
   // BODY (data max. 232 Byte, Array 0..231 of Byte) 
   IF #RD_WR = TRUE THEN
       // IO-Link write data record requested, copy data from "RECORD_IOL_DATA"
       #write.header.IOL.Control := B#16#02; // CONTROL B#16#02 = write data record
       #wrrec.length := INT_TO_UINT(#LEN) + UINT#8;  // data length header + data = IO-Link write data record
       #typeofrequest := 2; // write data record
       // copy IOL_RECORD_DATA in working area
       #i := INT#0;    // initialize loop counter 
       FOR #i := 0 TO #LEN - 1 DO
           #write.data[#i] := #RECORD_IOL_DATA[#i];
       END_FOR;
   ELSE
       // IO-Link read data record requested
       #write.header.IOL.Control := 16#03;  // CONTROL 16#03 = read data record
       #wrrec.length := UINT#8; // data length only header = IO-Link read data record
       #typeofrequest := 1; // read data record        
   END_IF;
   #sequencecontrol := 1;  // Start sequence
   ELSE
       ;
   END_IF;

   (*---------------------------------------------------------------------------------------------------------------------
               SEQUENCE CONTROL
   ---------------------------------------------------------------------------------------------------------------------*)
   CASE #sequencecontrol OF
       1:  // Check input parameter        
           IF #PORT < INT#0 OR #PORT > INT#63 THEN // PORT (Wrong port address = 0x8001)
               #ERROR := TRUE;
               #IOL_STATUS := DW#16#80010000;
               #sequencecontrol := 99; // aborting function with error
           ELSIF #IOL_INDEX < INT#0 OR #IOL_INDEX > INT#32767 THEN    // INDEX (Wrong index = 0x8002)
               #ERROR := TRUE;
               #IOL_STATUS := DW#16#80020000;
               #sequencecontrol := 99; // aborting function with error
           ELSIF #IOL_SUBINDEX < INT#0 OR #IOL_SUBINDEX > INT#255 THEN    // SUBINDEX (Wrong subindex = 0x8003)
               #ERROR := TRUE;
               #IOL_STATUS := DW#16#80030000;
               #sequencecontrol := 99; // aborting function with error
           ELSIF #typeofrequest = 2 AND (#LEN < 1 OR #LEN > 232) THEN  // LEN (wrong length for write data record = 0x8004)
               #ERROR := TRUE;
               #IOL_STATUS := DW#16#80050000;
               #sequencecontrol := 99; // aborting function with error
           ELSIF #typeofrequest = 1 AND (#LEN < 0 OR #LEN > 232) THEN  // LEN (wrong length for read data record = 0x8005)
               #ERROR := TRUE;
               #IOL_STATUS := DW#16#80060000;
               #sequencecontrol := 99; // aborting function with error
           ELSE    // all input parameter are right
               #sequencecontrol := 2;
           END_IF;

       2:  (*-------------------------------------------------------------------------------------------------------------
           WRREC = Write Data Record
           Note:
           To read data records, the IO-Link master modules needs to know which PORT is required. Therefore it is necessary
           to send at first a request via write data record (header, 8 byte). As response the IO-Link master module will 
           send the required data record.
           -------------------------------------------------------------------------------------------------------------*)
           #WRREC_Function(REQ := TRUE,
                           LEN := #wrrec.length,
                           DONE => #wrrec.done,
                           BUSY => #wrrec.busy,
                           ERROR => #wrrec.error,
                           STATUS => #wrrec.status,
                           RECORD := #write);
           // output status during write data record
           IF #wrrec.busy THEN
               #STATUS := #wrrec.status;
               #IOL_STATUS := DW#16#00020000;  // 0002 = writing in progress 
           ELSIF #wrrec.error THEN
               #tmpDWORD := #wrrec.status AND DW#16#00FFFF00;  // filter status
               IF #tmpDWORD = DW#16#0080C200 THEN    // if resource #BUSY (#STATUS=80C2), then ... 
                   #sequencecontrol := 3;  // ... repeat write data record
               ELSE
                   #ERROR := TRUE;
                   #STATUS := #wrrec.status;   // ... otherwise output error status of "WRREC"
                   #IOL_STATUS := DW#16#80530000;  // ... with note '8053' = error status of "WRREC"
                   #sequencecontrol := 99; // aborting function with error
               END_IF;
           ELSIF #wrrec.done = TRUE THEN   // wait for write data record finish without error
               #TP_poll(IN := TRUE,
                        PT := T#100ms);    // poll for response
               #sequencecontrol := 4;
           ELSE
               ;
           END_IF;

       3:  // repeat write data record because resource was busy
           #WRREC_Function(REQ := FALSE);
           #sequencecontrol := 2;

       4:  // wait and poll for response = Read Data Record (RDREC)
           #WRREC_Function(REQ := FALSE);
           #TP_poll(IN := TRUE,
                    PT := T#100ms);

           // if poll rate executed then start read data record (on falling edge)
           #F_TRIG_poll := #TP_poll.Q = FALSE AND #F_TRIG_poll_old = TRUE;
           #F_TRIG_poll_old := #TP_poll.Q = TRUE;

           // RDREC = Read Data Record
           #RDREC_Function(REQ := #F_TRIG_poll,
                           MLEN := UINT#0, // length = 0 = read all data which are available
                           VALID => #rdrec.valid,
                           BUSY => #rdrec.busy,
                           ERROR => #rdrec.error,
                           STATUS => #rdrec.status,
                           LEN => #rdrec.length,
                           RECORD := #read);
           // output status during read data record
           IF #rdrec.busy THEN
               #STATUS := #rdrec.status;
               #IOL_STATUS := DW#16#00030000; // 16#0003 = reading in progress
           ELSIF #rdrec.error = TRUE THEN
               #tmpDWORD := #rdrec.status AND DW#16#00FFFF00;  // filter status
               IF #tmpDWORD = DW#16#0080C200 THEN  // if resource busy (status=80C2), then ... 
                   #sequencecontrol := 5;  // ... repeat read data record / continue polling
               ELSE
                   #ERROR := TRUE;
                   #STATUS := #rdrec.status;   // ... otherwise output error code of "RDREC"
                   #IOL_STATUS := DW#16#80520000;  // ... with note '8052' = error status of "RDREC"
                   #sequencecontrol := 99; // aborting function with error
               END_IF;
           ELSIF #rdrec.valid THEN
               IF  // check the response wether it matches the request (compare PORT, INDEX and SUBINDEX)
                   (#write.header.CALL.Port <> #read.header.CALL.Port) OR
                   (#write.header.IOL.Index_HighByte <> #read.header.IOL.Index_HighByte) OR
                   (#write.header.IOL.Index_LowByte <> #read.header.IOL.Index_LowByte) OR
                   (#write.header.IOL.Subindex <> #read.header.IOL.Subindex)
               THEN    // read data record don't match the request
                   #ERROR := TRUE;
                   #STATUS := #rdrec.status;
                   #IOL_STATUS := DW#16#70000000;  // output status '7000', no consistent data
                   #sequencecontrol := 99; // aborting function with error
               ELSIF #read.header.IOL.Control = B#16#80 THEN   // check the response for IO-Link errors
                   // State 0x80 = IOL_CALL_RES PDU shows IO-Link error detect
                   #ERROR := TRUE;
                   #STATUS := DW#16#00000000;
                   #IOL_STATUS.%B3 := #read.data[0];   // IO-Link master error code
                   #IOL_STATUS.%B2 := #read.data[1];   // IO-Link master error code
                   #IOL_STATUS.%B1 := #read.data[2];  // IO-Link device error code
                   #IOL_STATUS.%B0 := #read.data[3];  // IO-Link device additional error code

                   #sequencecontrol := 99; // aborting function with error
               ELSE    // read data are valid = output
                   #DONE_VALID := TRUE;
                   #BUSY := FALSE;
                   #ERROR := FALSE;
                   #STATUS := DW#16#00000000;
                   #IOL_STATUS := DW#16#00000000;  // request finished

                   IF #typeofrequest = 1 THEN
                       #RD_LEN := UINT_TO_INT(#rdrec.length - UINT#8);  // device parameter cover header and data,
                       // only data will be output
                       #i := INT#0; // initialize loop counter
                       FOR #i := 0 TO UINT_TO_INT(#rdrec.length - UINT#8 - UINT#1) DO
                           #RECORD_IOL_DATA[#i] := #read.data[#i];
                       END_FOR;
                   ELSE
                       ;
                   END_IF;
                   #sequencecontrol := 98;
               END_IF;
           ELSE
               ;
           END_IF;

       5:  // poll again for response because resource was busy
           #TP_poll(IN := FALSE,
                    PT := T#100ms);
           #RDREC_Function(REQ := FALSE,
                           RECORD := #read);
           #sequencecontrol := 4;  // ... repeat read data record / continue polling   

       98: // request done successfully
           #TP_poll(IN := FALSE,
                    PT := T#100ms);
           #RDREC_Function(REQ := FALSE,
                           RECORD := #read);
           IF #REQ = FALSE THEN
               #DONE_VALID := FALSE;
               #BUSY := FALSE;
               #ERROR := FALSE;
               #RD_LEN := INT#0;
               #STATUS := DW#16#00000000;
               #IOL_STATUS := DW#16#00010000; // ready for new request
               #sequencecontrol := 0;
               #typeofrequest := 0;
           ELSE
               ;
           END_IF;

       99: // Function aborted with error
           #TP_poll(IN := FALSE,
                    PT := T#100ms);
           #WRREC_Function(REQ := FALSE);
           #RDREC_Function(REQ := FALSE,
                           RECORD := #read);
           #DONE_VALID := FALSE;
           #BUSY := FALSE;
           #RD_LEN := INT#0;
           #sequencecontrol := 0;
           #typeofrequest := 0;

       ELSE  // no relevant case, ready for new request
           #WRREC_Function(REQ := FALSE);
           #RDREC_Function(REQ := FALSE,
                           RECORD := #read);
           #TP_poll(IN := FALSE,
                    PT := T#100ms);
           #TON_monitoring(IN := FALSE,
                           PT := T#20s);
           #sequencecontrol := 0;
           #typeofrequest := 0;
   END_CASE;

   (*---------------------------------------------------------------------------------------------------------------------
               MONITORING
   ---------------------------------------------------------------------------------------------------------------------*)
   #TON_monitoring(IN := #sequencecontrol > 0 AND #sequencecontrol < 98,
                   PT := T#20s);
   IF #TON_monitoring.Q THEN
       #ERROR := TRUE;
       #IOL_STATUS := DW#16#80000000; // request time out       
       #sequencecontrol := 99; // aborting function with error
   END_IF;
END_FUNCTION_BLOCK

(* ===== HMI "HMI_RT_1" =====
system functions are stored by id; their names below are inferred from use
connection "HMI_Connection_1": ETHERNET, SMART_S7_1200_OMS

HMI tags "Default tag table"
   "Emergency Stop Stacker" : Bool = PLC 113S1 AT %I1.0, 1 s
   "Avarie Conveior 4 stacker" : Bool = PLC 128U1_Fault AT %I5.1, 1 s
   "Prezenta aer" : Bool = PLC 151S1 AT %I2.0, 1 s
   "Protectie cuplata Conveior 1 alimentare destacker" : Bool = PLC 120Q1 AT %I2.2, 1 s
   "Protectie cuplata Conveior 2 iesire destacker" : Bool = PLC 122Q1 AT %I2.7, 1 s
   "Avarie Conveior 1 alimentare destacker" : Bool = PLC 120U1_Fault AT %I2.6, 1 s
   "Avarie Conveior 2 iesire destacker" : Bool = PLC 122U1_Fault AT %I3.3, 1 s
   "Contactor cuplat Conveior 1 alimentare destacker" : Bool = PLC 121K1 AT %I2.3, 1 s
   "Contactor cuplat Conveior 2 iesire destacker" : Bool = PLC 123K1 AT %I3.0, 1 s
   "Frana decuplata Conveior 1 alimentare destacker" : Bool = PLC 120K1 AT %I2.4, 1 s
   "Frana decuplata Conveior 2 iesire destacker" : Bool = PLC 122K1 AT %I3.1, 1 s
   "Functionare Conveior 1 alimentare destacker" : Bool = PLC 120U1_PowerOK AT %I2.5, 1 s
   "Functionare Conveior 2 iesire destacker" : Bool = PLC 122U1_PowerOK AT %I3.2, 1 s
   "Senzor 1 proximitate softstarter aer destacker" : Bool = PLC 142VFA1_SQ1 AT %I6.4, 1 s
   "Senzor 2 proximitate softstarter aer destacker" : Bool = PLC 142VFA1_SQ2 AT %I6.5, 1 s
   "Reset safety Destacker" : Bool = PLC 1XXS2 AT %I68.6, 1 s
   "Comanda 1 softstarter aer destacker" : Bool = PLC "Comanda 1 softstarter aer stacker_new" AT %Q64.1, 1 s
   "Cuplare contactor VFD Conveior 1 alimentare destacker" : Bool = PLC CSN3_PowerOK AT %Q7.3, 1 s
   "Fault Aknowledge VFD Conveior 1 alimentare destacker" : Bool = PLC CSN3_FaultAck AT %Q10.0, 1 s
   "ON/OFF1 VFD Conveior 1 alimentare destacker" : Bool = PLC CSN3_Start AT %Q7.4, 1 s
   "Cuplare contactor VFD Conveior 2 iesire destacker" : Bool = PLC CSN4_PowerOK AT %Q7.5, 1 s
   "Fault Aknowledge VFD Conveior 2 iesire destacker" : Bool = PLC CSN4_FaultAck AT %Q10.1, 1 s
   "ON/OFF1 VFD Conveior 2 iesire destacker" : Bool = PLC CSN4_Start AT %Q7.6, 1 s
   "Contactor cuplat Conveior 4 descarcare stacker" : Bool = PLC 129K1 AT %I4.6, 1 s
   "Frana decuplata Conveior 4 descarcare stacker" : Bool = PLC 128K1 AT %I4.7, 1 s
   "Functionare Conveior 4 stacker" : Bool = PLC 128U1_PowerOK AT %I5.0, 1 s
   "Protectie cuplata Conveior 4 descarcare stacker" : Bool = PLC 128Q1 AT %I4.5, 1 s
   "Cuplare contactor VFD Conveior 4 descarcare stacker" : Bool = PLC CS4_PowerOK AT %Q8.5, 1 s
   "Fault Aknowledge VFD Conveior 4 descarcare stacker" : Bool = PLC CS4_FaultAck AT %Q10.3, 1 s
   "ON/OFF1 VFD Conveior 4 descarcare stacker" : Bool = PLC CS4_Start AT %Q8.6, 1 s
   "Avarie Conveior 3 transfer palet 2" : Bool = PLC 126U1_Fault AT %I4.4, 1 s
   "Contactor cuplat Conveior 3 transfer palet 2" : Bool = PLC 127K1 AT %I4.1, 1 s
   "Frana decuplata Conveior 3 transfer palet 2" : Bool = PLC 126K1 AT %I4.2, 1 s
   "Functionare Conveior 1 preluare paleti OK" : Bool = PLC 124K1 AT %I3.5, 1 s
   "Functionare Conveior 2 transfer palet 1" : Bool = PLC 125K1 AT %I3.7, 1 s
   "Functionare Conveior 3 transfer palet 2" : Bool = PLC 126U1_PowerOK AT %I4.3, 1 s
   "Protectie cuplata Conveior 1 preluare paleti OK" : Bool = PLC 124Q1 AT %I3.4, 1 s
   "Protectie cuplata Conveior 2 transfer palet 1" : Bool = PLC 125Q1 AT %I3.6, 1 s
   "Protectie cuplata Conveior 3 transfer palet 2" : Bool = PLC 126Q1 AT %I4.0, 1 s
   "Cuplare contactor VFD Conveior 3 transfer palet 2" : Bool = PLC CS3_PowerOK AT %Q8.3, 1 s
   "Fault Aknowledge VFD Conveior 3 transfer palet 2" : Bool = PLC CS3_FaultAck AT %Q10.2, 1 s
   "ON/OFF1 VFD Conveior 3 transfer palet 2" : Bool = PLC CS3_Start AT %Q8.4, 1 s
   "Softstarter aer 1.1 Conveior 1 preluare paleti OK" : Bool = PLC "Softstarter aer 1.1 Conveior 1 preluare paleti OK" AT %Q8.1, 1 s
   "Softstarter aer 1.2 Conveior 1 preluare paleti OK" : Bool = PLC "Softstarter aer 1.2 Conveior 1 preluare paleti OK" AT %Q8.2, 1 s
   "Start Conveior 1 preluare paleti OK" : Bool = PLC CS1_Start AT %Q8.0, 1 s
   "Start Conveior 2 transfer palet 1" : Bool = PLC CS2_Start AT %Q7.0, 1 s
   "Comanda 2 softstarter aer destacker" : Bool = PLC "Comanda 2 softstarter aer stacker_new" AT %Q66.1, 1 s
   "Comanda 1 softstarter aer stacker" : Bool = PLC "Comanda 1 softstarter aer stacker" AT %Q72.1, 1 s
   "Comanda 2 softstarter aer stacker" : Bool = PLC "Comanda 2 softstarter aer stacker" AT %Q74.1, 1 s
   "MD_IS1_SC_X1.0" : Bool = PLC "MD_IS1_SC_X1.0" AT %I70.0, 1 s
   "MD_IS1_SC_X1.1" : Bool = PLC "MD_IS1_SC_X1.1" AT %I70.1, 1 s
   "MD_IS1_SC_X1.2" : Bool = PLC "MD_IS1_SC_X1.2" AT %I70.2, 1 s
   "MD_IS1_SC_X1.3" : Bool = PLC "MD_IS1_SC_X1.3" AT %I70.3, 1 s
   "MD_IS1_SC_X1.4" : Bool = PLC "MD_IS1_SC_X1.4" AT %I70.4, 1 s
   "MD_IS1_SC_X1.5" : Bool = PLC "MD_IS1_SC_X1.5" AT %I70.5, 1 s
   "MD_IS1_SC_X1.6" : Bool = PLC "MD_IS1_SC_X1.6" AT %I70.6, 1 s
   "MD_IS1_SC_X1.7" : Bool = PLC "MD_IS1_SC_X1.7" AT %I70.7, 1 s
   "MD_IS2_SC_X1.0" : Bool = PLC "MD_IS2_SC_X1.0" AT %I75.0, 1 s
   "MD_IS2_SC_X1.1" : Bool = PLC "MD_IS2_SC_X1.1" AT %I75.1, 1 s
   "MD_IS2_SC_X1.2" : Bool = PLC "MD_IS2_SC_X1.2" AT %I75.2, 1 s
   "MD_IS2_SC_X1.3" : Bool = PLC "MD_IS2_SC_X1.3" AT %I75.3, 1 s
   "MD_IS2_SC_X1.4" : Bool = PLC "MD_IS2_SC_X1.4" AT %I75.4, 1 s
   "MD_IS2_SC_X1.5" : Bool = PLC "MD_IS2_SC_X1.5" AT %I75.5, 1 s
   "MD_IS2_SC_X1.6" : Bool = PLC "MD_IS2_SC_X1.6" AT %I75.6, 1 s
   "MD_IS2_SC_X1.7" : Bool = PLC "MD_IS2_SC_X1.7" AT %I75.7, 1 s
   "MD_OS_SC_X1.0" : Bool = PLC "MD_OS_SC_X1.0" AT %I92.0, 1 s
   "MD_OS_SC_X1.1" : Bool = PLC "MD_OS_SC_X1.1" AT %I93.0, 1 s
   "MD_OS_SC_X1.2" : Bool = PLC "MD_OS_SC_X1.2" AT %I92.1, 1 s
   "MD_OS_SC_X1.3" : Bool = PLC "MD_OS_SC_X1.3" AT %I93.1, 1 s
   "MD_OS_SC_X1.4" : Bool = PLC "MD_OS_SC_X1.4" AT %I92.2, 1 s
   "MD_OS_SC_X1.5" : Bool = PLC "MD_OS_SC_X1.5" AT %I93.2, 1 s
   "MS_IS1_SC_X1.0" : Bool = PLC "MS_IS1_SC_X1.0" AT %I80.0, 1 s
   "MS_IS1_SC_X1.1" : Bool = PLC "MS_IS1_SC_X1.1" AT %I80.1, 1 s
   "MS_IS1_SC_X1.2" : Bool = PLC "MS_IS1_SC_X1.2" AT %I80.2, 1 s
   "MS_IS1_SC_X1.3" : Bool = PLC "MS_IS1_SC_X1.3" AT %I80.3, 1 s
   "MS_IS1_SC_X1.4" : Bool = PLC "MS_IS1_SC_X1.4" AT %I80.4, 1 s
   "MS_IS1_SC_X1.5" : Bool = PLC "MS_IS1_SC_X1.5" AT %I80.5, 1 s
   "MS_IS1_SC_X1.6" : Bool = PLC "MS_IS1_SC_X1.6" AT %I80.6, 1 s
   "MS_IS1_SC_X1.7" : Bool = PLC "MS_IS1_SC_X1.7" AT %I80.7, 1 s
   "MS_IS2_SC_X1.0" : Bool = PLC "MS_IS2_SC_X1.0" AT %I85.0, 1 s
   "MS_IS2_SC_X1.1" : Bool = PLC "MS_IS2_SC_X1.1" AT %I85.1, 1 s
   "MS_IS2_SC_X1.2" : Bool = PLC "MS_IS2_SC_X1.2" AT %I85.2, 1 s
   "MS_IS2_SC_X1.3" : Bool = PLC "MS_IS2_SC_X1.3" AT %I85.3, 1 s
   "MS_IS2_SC_X1.4" : Bool = PLC "MS_IS2_SC_X1.4" AT %I85.4, 1 s
   "MS_IS2_SC_X1.5" : Bool = PLC "MS_IS2_SC_X1.5" AT %I85.5, 1 s
   "MS_IS2_SC_X1.6" : Bool = PLC "MS_IS2_SC_X1.6" AT %I85.6, 1 s
   "MS_IS2_SC_X1.7" : Bool = PLC "MS_IS2_SC_X1.7" AT %I85.7, 1 s
   "MS_OS_SC_X1.0" : Bool = PLC "MS_OS_SC_X1.0" AT %I101.0, 1 s
   "MS_OS_SC_X1.1" : Bool = PLC "MS_OS_SC_X1.1" AT %I102.0, 1 s
   "MS_OS_SC_X1.2" : Bool = PLC "MS_OS_SC_X1.2" AT %I101.1, 1 s
   "MS_OS_SC_X1.3" : Bool = PLC "MS_OS_SC_X1.3" AT %I102.1, 1 s
   "MS_OS_SC_X1.4" : Bool = PLC "MS_OS_SC_X1.4" AT %I101.2, 1 s
   "MS_OS_SC_X1.5" : Bool = PLC "MS_OS_SC_X1.5" AT %I102.2, 1 s
   "DS_Comanda cilindru vertical jos" : Bool = PLC "SN_Comanda cilindru vertical jos" AT %Q66.0, 1 s
   "DS_Comanda cilindru vertical sus" : Bool = PLC "SN_Comanda cilindru vertical sus" AT %Q64.0, 1 s
   "DS_Comanda furca retrasa" : Bool = PLC "SN_Comanda furca retrasa" AT %Q65.0, 1 s
   "DB_PalletDispenser_PD2_De_Stacking_DB_PD1_MiddlePosition" : Bool = PLC DB_PalletDispenser_PD2_Stacking_New_DB.PD1.MiddlePosition, 1 s
   "DB_PalletDispenser_PD2_De_Stacking_DB_PD1_Up" : Bool = PLC DB_PalletDispenser_PD2_Stacking_New_DB.PD1.Up, 1 s
   "DB_PalletDispenser_PD2_De_Stacking_DB_PD1_Down" : Bool = PLC DB3_FAULTS.Alarm_Safety_S, 1 s
   "DB_PalletDispenser_PD2_De_Stacking_DB_PD1_Forks_In" : Bool = PLC DB3_FAULTS.Alarm_Safety_Z2, 1 s
   "DB_PalletDispenser_PD2_De_Stacking_DB_PD1_Forks_Out" : Bool = PLC DB_PalletDispenser_PD2_Stacking_New_DB.PD1.Forks_Out, 1 s
   "DB_PalletDispenser_PD2_De_Stacking_DB_Alarm_Active" : Bool = PLC DB3_FAULTS.Alarm_CD1, 1 s
   "DB_PalletDispenser_PD2_Stacking_DB_PD1_MiddlePosition" : Bool = PLC DB_PalletDispenser_PD2_Stacking_DB.PD1.MiddlePosition, 1 s
   "DB_PalletDispenser_PD2_Stacking_DB_PD1_Up" : Bool = PLC DB_PalletDispenser_PD2_Stacking_DB.PD1.Up, 1 s
   "DB_PalletDispenser_PD2_Stacking_DB_PD1_Down" : Bool = PLC DB_PalletDispenser_PD2_Stacking_DB.PD1.Down, 1 s
   "DB_PalletDispenser_PD2_Stacking_DB_PD1_Forks_In" : Bool = PLC DB_PalletDispenser_PD2_Stacking_DB.PD1.Forks_In, 1 s
   "DB_PalletDispenser_PD2_Stacking_DB_PD1_Forks_Out" : Bool = PLC DB_PalletDispenser_PD2_Stacking_DB.PD1.Forks_Out, 1 s
   "DB_PalletDispenser_PD2_Stacking_DB_Alarm_Active" : Bool = PLC DB_PalletDispenser_PD2_Stacking_DB.Alarm.Active, 1 s
   "S_Comanda cilindru vertical jos" : Bool = PLC "S_Comanda cilindru vertical jos" AT %Q74.0, 1 s
   "S_Comanda cilindru vertical sus" : Bool = PLC "S_Comanda cilindru vertical sus" AT %Q72.0, 1 s
   "S_Comanda furca retrasa" : Bool = PLC "S_Comanda furca retrasa" AT %Q73.0, 1 s
   "S_Comanda furca extinsa" : Bool = PLC "S_Comanda furca extinsa" AT %Q75.0, 1 s
   "Destacker 110KF1 Safety Relay" : Bool = PLC 110KF1 AT %I0.0, 1 s
   "Destacker 111KF1 Safety Barrier Relay" : Bool = PLC 111KF1 AT %I0.1, 1 s
   "Emergency Stop Destacker" : Bool = PLC 110S1 AT %I0.6, 1 s
   "Emergency Stop Zone 2" : Bool = PLC 112S1 AT %I0.7, 1 s
   "Stacker 113KF1 Safety Relay" : Bool = PLC 113KF1 AT %I0.3, 1 s
   "Stacker 114KF1 Safety Barrier Relay 1" : Bool = PLC 114KF1 AT %I0.4, 1 s
   "Stacker 115KF1 Safety Barrier Relay 2" : Bool = PLC 115KF1 AT %I0.5, 1 s
   "Zone 2 112KF1 Safety Relay" : Bool = PLC 112KF1 AT %I0.2, 1 s
   "Reset Destacker 110KF1 Safety Relay" : Bool = PLC 153K1 AT %Q0.0, 1 s
   "Reset Destacker 111KF1 Safety Barrier Relay" : Bool = PLC 153K2 AT %Q0.1, 1 s
   "Reset safety Zone 2" : Bool = PLC 155S1 AT %I1.1, 1 s
   "Reset Stacker 113KF1 Safety Relay" : Bool = PLC 153K4 AT %Q0.3, 1 s
   "Reset Stacker 114KF1 Safety Barrier Relay 1" : Bool = PLC 153K5 AT %Q0.4, 1 s
   "Reset Stacker 115KF1 Safety Barrier Relay 2" : Bool = PLC 153K6 AT %Q0.5, 1 s
   "Reset Zone 2 112KF1 Safety Relay" : Bool = PLC 153K3 AT %Q0.2, 1 s
   "FB_AlarmCounter_DB_Counters_Destacker 110KF1 Safety Relay_CV" : Int = PLC FB_AlarmCounter_DB.Counters."Destacker 110KF1 Safety Relay".CV, 1 s
   "FB_AlarmCounter_DB_Counters_Destacker 111KF1 Safety Barrier Relay_CV" : Int = PLC FB_AlarmCounter_DB.Counters."Destacker 111KF1 Safety Barrier Relay".CV, 1 s
   "FB_AlarmCounter_DB_Counters_Zone 2 112KF1 Safety Relay_CV" : Int = PLC FB_AlarmCounter_DB.Counters."Zone 2 112KF1 Safety Relay".CV, 1 s
   "FB_AlarmCounter_DB_Counters_Stacker 113KF1 Safety Relay_CV" : Int = PLC FB_AlarmCounter_DB.Counters."Stacker 113KF1 Safety Relay".CV, 1 s
   "FB_AlarmCounter_DB_Counters_Stacker 114KF1 Safety Barrier Relay 1_CV" : Int = PLC FB_AlarmCounter_DB.Counters."Stacker 114KF1 Safety Barrier Relay 1".CV, 1 s
   "FB_AlarmCounter_DB_Counters_Stacker 115KF1 Safety Barrier Relay 2_CV" : Int = PLC FB_AlarmCounter_DB.Counters."Stacker 115KF1 Safety Barrier Relay 2".CV, 1 s
   "FB_AlarmCounter_DB_Counters_Emergency Stop Destacker_CV" : Int = PLC FB_AlarmCounter_DB.Counters."Emergency Stop Destacker".CV, 1 s
   "FB_AlarmCounter_DB_Counters_Emergency Stop Zone 2_CV" : Int = PLC FB_AlarmCounter_DB.Counters."Emergency Stop Zone 2".CV, 1 s
   "FB_AlarmCounter_DB_Counters_Emergency Stop Stacker_CV" : Int = PLC FB_AlarmCounter_DB.Counters."Emergency Stop Stacker".CV, 1 s
   "FB_EnergyCounter_DB_Counters_LastHour_CV" : UInt = PLC FB_EnergyCounter_DB.Counters.LastHour.CV, 1 s
   "FB_EnergyCounter_DB_Counters_LastDay_CV" : UDInt = PLC FB_EnergyCounter_DB.Counters.LastDay.CV, 1 s
   "FB_EnergyCounter_DB_Counters_LastMonth_CV" : UDInt = PLC FB_EnergyCounter_DB.Counters.LastMonth.CV, 1 s
   "Aliniere palet" : Bool = PLC CSN1_SQ3 AT %I68.1, 1 s
   "Centror extins" : Bool = PLC CP2_SQ3 AT %I79.5, 1 s
   "Centror retras" : Bool = PLC CP2_SQ2 AT %I78.5, 1 s
   "Detectie 1 aliniament palet" : Bool = PLC "Detectie 1 aliniament palet" AT %I69.1, 1 s
   "Detectie 2 aliniament palet" : Bool = PLC "Detectie 2 aliniament palet" AT %I68.2, 1 s
   "Detectie palet" : Bool = PLC "SN_Detectie palet" AT %I73.4, 1 s
   "DS_Cilindru extins" : Bool = PLC "SN_Cilindru extins" AT %I74.6, 1 s
   "DS_Cilindru retras" : Bool = PLC "SN_Cilindru retras" AT %I74.1, 1 s
   "DS_Cilindru vertical jos" : Bool = PLC "SN_Cilindru vertical jos" AT %I73.5, 1 s
   "DS_Cilindru vertical mijloc" : Bool = PLC "SN_Cilindru vertical mijloc" AT %I73.3, 1 s
   "DS_Cilindru vertical sus" : Bool = PLC "SN_Cilindru vertical sus" AT %I73.2, 1 s
   "DS_Lungime 1" : Bool = PLC CSN3_SQ2 AT %I68.3, 1 s
   "DS_Lungime 2" : Bool = PLC CSN3_SQ3 AT %I69.3, 1 s
   "DS_Lungime 3" : Bool = PLC CSN4_SQ1 AT %I68.4, 1 s
   "Feed palet" : Bool = PLC SN_Prez_conveyor_volum AT %I69.6, 1 s
   "Inaltime maxima" : Bool = PLC "Inaltime maxima" AT %I69.0, 1 s
   "Masurare lungime" : Bool = PLC CS2_SQ1 AT %I78.2, 1 s
   "Prezenta palet iesire" : Bool = PLC SN_Switch_Iesire AT %I69.4, 1 s
   "Prezenta palet_capat_conveyor" : Bool = PLC CS1_SQ3 AT %I78.1, 1 s
   "Prezenta palet_centror" : Bool = PLC "S_Prezenta palet_centror" AT %I79.1, 1 s
   "Prezenta palet_dreapta" : Bool = PLC "Prezenta palet_dreapta" AT %I79.0, 1 s
   "Prezenta palet_stanga" : Bool = PLC CS1_SQ1 AT %I78.0, 1 s
   "Prezenta_stiva" : Bool = PLC CS4_SQ1 AT %I78.4, 1 s
   "Prezenta stiva" : Bool = PLC CSN1_SQ1 AT %I68.0, 1 s
   "Protectie cuplata Circular masa fixa" : Bool = PLC 104F1 AT %I5.4, 1 s
   "Protectie cuplata HMI" : Bool = PLC 149F1 AT %I7.0, 1 s
   "Protectie cuplata Iluminat" : Bool = PLC 105F2 AT %I2.1, 1 s
   "Protectie cuplata Masina demontare paleti dreapta" : Bool = PLC 103F1 AT %I5.3, 1 s
   "Protectie cuplata Masina demontare paleti stanga" : Bool = PLC 102F1 AT %I5.2, 1 s
   "Protectie cuplata Post reparatie stanga+dreapta" : Bool = PLC 105F1 AT %I5.5, 1 s
   "Protectie cuplata Post reparatii minore" : Bool = PLC 106F1 AT %I5.6, 1 s
   "Protectie cuplata TELE" : Bool = PLC 107F1 AT %I5.7, 1 s
   "S_Cilindru extins" : Bool = PLC "S_Cilindru extins" AT %I84.6, 1 s
   "S_Cilindru retras" : Bool = PLC "S_Cilindru retras" AT %I84.1, 1 s
   "S_Cilindru vertical jos" : Bool = PLC "S_Cilindru vertical jos" AT %I83.5, 1 s
   "S_Cilindru vertical mijloc" : Bool = PLC "S_Cilindru vertical mijloc" AT %I83.3, 1 s
   "S_Cilindru vertical sus" : Bool = PLC "S_Cilindru vertical sus" AT %I83.2, 1 s
   "S_Lungime 1" : Bool = PLC CS3_SQ1 AT %I79.2, 1 s
   "S_Lungime 2" : Bool = PLC CS3_SQ2 AT %I78.3, 1 s
   "S_Lungime 3" : Bool = PLC CS3_SQ3 AT %I79.3, 1 s
   "S_Detectie palet" : Bool = PLC "S_Detectie palet" AT %I83.4, 1 s
   "Senzor 1 prezenta stiva" : Bool = PLC "Senzor 1 prezenta stiva" AT %I68.5, 1 s
   "Senzor 1 proximitate softstarter aer stacker" : Bool = PLC 143VFA1_SQ1 AT %I83.7, 1 s
   "Senzor 1 proximitate softstarter aer zona 2" : Bool = PLC 141VFA1_SQ1 AT %I7.1, 1 s
   "Senzor 2 prezenta stiva" : Bool = PLC "Senzor 2 prezenta stiva" AT %I69.5, 1 s
   "Senzor 2 proximitate softstarter aer stacker" : Bool = PLC 143VFA1_SQ2 AT %I84.7, 1 s
   "Senzor 2 proximitate softstarter aer zona 2" : Bool = PLC 141VFA1_SQ2 AT %I7.2, 1 s
   "Senzor destacking" : Bool = PLC "SN_Senzor stacking" AT %I73.1, 1 s
   "Senzor stacking" : Bool = PLC "S_Senzor stacking" AT %I83.1, 1 s
   "Start masurare lungime" : Bool = PLC CSN3_SQ1 AT %I69.2, 1 s
   "DS_Comanda furca extinsa" : Bool = PLC "SN_Comanda furca extinsa" AT %Q67.0, 1 s
   "DB20_DATA_HMI_Step_Destacker" : Int = PLC DB20_DATA_HMI.Step_Destacker, 1 s
   "DB20_DATA_HMI_Step_Stacker" : Int = PLC DB20_DATA_HMI.Step_Stacker, 1 s
   "Maintenance" : Bool = PLC Maintenance AT %M5.0, 1 s
   "Rez_G7_DS" : Bool = PLC Rez_G7_DS AT %M6.0, 1 s
   "Rez_G7_S" : Bool = PLC Rez_G7_S AT %M6.1, 1 s
   "Fault_Length_DS" : Bool = PLC Fault_Length_DS AT %M6.2, 1 s
   "Fault_Length_DS_ACK" : Bool = PLC Fault_Length_DS_ACK AT %M6.4, 1 s
   "Length_DS_HMI_1" : Bool = PLC Length_DS_HMI_1 AT %M14.0, 1 s
   "Length_DS_HMI_2" : Bool = PLC Length_DS_HMI_2 AT %M14.1, 1 s
   "Length_DS_HMI_3" : Bool = PLC Length_DS_HMI_3 AT %M14.2, 1 s
   "Length_S_HMI_1" : Bool = PLC Length_S_HMI_1 AT %M14.3, 1 s
   "Length_S_HMI_2" : Bool = PLC Length_S_HMI_2 AT %M14.4, 1 s
   "Length_S_HMI_3" : Bool = PLC Length_S_HMI_3 AT %M14.5, 1 s
   "Fault_Length_S_ACK" : Bool = PLC Fault_Length_S_ACK AT %M6.5, 1 s
   "Fault_Length_S" : Bool = PLC Fault_Length_S AT %M6.3, 1 s
   "DB_MDM_SN_step" : USInt = PLC O.Centror_A.AlarmW, 1 s
   "DB_MDM_S_step" : USInt = PLC DB3_FAULTS.Alarm_CD2, 1 s
   "s_f{1}_step" : USInt = PLC s.f[5].AlarmW, 1 s
   "s_f{1}_almt" : Bool = PLC s.f[4].AlarmW, 1 s
   "s_f{3}_step" : USInt = PLC s.f[3].AlarmW, 1 s
   "s_f{4}_step" : USInt = PLC s.f[2].AlarmW, 1 s
   "s_f{5}_step" : USInt = PLC FB_ProductionStatistics_DB.Counters.Destroyed.LastDay.CV, 1 s
   "s_f{3}_almt" : Bool = PLC FB_ProductionStatistics_DB.Counters.Repairs.LastDay.CV, 1 s
   "s_f{4}_almt" : Bool = PLC "Manual_Comanda 1 softstarter aer destacker", 1 s
   "s_f{5}_almt" : Bool = PLC "Manual_Comanda 2 softstarter aer destacker", 1 s
   "sn_f{2}_step" : USInt = PLC O.CilindruVerticalStacker.ButRet, 1 s
   "sn_f{3}_step" : USInt = PLC O.CilindruVerticalStacker.ButAv, 1 s
   "sn_f{4}_step" : USInt = PLC O.FurcaStacker.ButAv, 1 s
   "sn_f{5}_step" : USInt = PLC O.FurcaStacker.ButRet, 1 s
   "sn_f{2}_almt" : Bool = PLC "Manual_Cuplare contactor VFD Conveior 1 alimentare destacker", 1 s
   "sn_f{3}_almt" : Bool = PLC "Manual_Fault Aknowledge VFD Conveior 1 alimentare destacker", 1 s
   "sn_f{4}_almt" : Bool = PLC "Manual_ON/OFF1 VFD Conveior 1 alimentare destacker", 1 s
   "sn_f{5}_almt" : Bool = PLC "Manual_Cuplare contactor VFD Conveior 2 iesire destacker", 1 s
   "sn_f{1}_almt" : Bool = PLC "Manual_ON/OFF1 VFD Conveior 2 iesire destacker", 1 s
   "sn_f{1}_step" : USInt = PLC "Manual_Reset Destacker 110KF1 Safety Relay", 1 s
   "s_f{2}_step" : USInt = PLC "Manual_Reset Destacker 111KF1 Safety Barrier Relay", 1 s
   "s_f{2}_almt" : Bool = PLC "Manual_Reset Zone 2 112KF1 Safety Relay", 1 s

HMI tags "Alarms"
   "DS_AlarmMovement" : Word = PLC DS_AlarmMovement AT %MW2, 1 s
   "S_AlarmMovement" : Word = PLC S_AlarmMovement AT %MW4, 1 s

HMI tags "UserManagement"
   "CurrentUser" : WString[254], internal
   "CurrentUserGroup" : Int, internal

HMI tags "Statistics"
   "PalletsLastMonth" : Int, internal
   "PalletsLastWeek" : Int, internal
   "PalletsPerShift" : Array [0..8] of Int, internal

HMI tags "UI"
   "CurrentScreenStatistics" : Int, internal
   "CurrentScreenManual" : Bool = PLC DB20_DATA_HMI.Maintenance, 1 s
   "SwitchTestBit" : Bool, internal

discrete alarms
   1: 'Alarma destacker miscare verticala', class Errors, trigger "DS_AlarmMovement" bit 0
   2: 'Alarma destacker miscare furci', class Errors, trigger "DS_AlarmMovement" bit 1
   3: 'Alarma destacker pozitie', class Errors, trigger "DS_AlarmMovement" bit 2
   4: 'Alarma stacker miscare verticala', class Errors, trigger "S_AlarmMovement" bit 0
   5: 'Alarma stacker miscare furci', class Errors, trigger "S_AlarmMovement" bit 1
   6: 'Alarma stacker pozitie', class Errors, trigger "S_AlarmMovement" bit 2

text list "Text_list_1": 0 'Yes / Da'; 1 'No / Nu'

graphic list "@DiagnosticsStates": 0 '@Diagnostics_StateGood'; 1 '@Diagnostics_StateBad'

graphic list "List": 1 'Graphic_4'; 2 'Graphic_6'; 4..16 'Graphic_7'

screen "Main" 800x480, template "TemplateWithClock"
   Button "Button_1" at 8,392 size 136x80; TextOn 'Pagina Principala'; TextOff 'Pagina Principala'
      on Press: ActivateScreen("Main", 0)
   Button "Button_2" at 152,392 size 136x80; TextOff 'Mod Manual'; Authorization "Operate"
      on Press: ActivateScreen("Manual.General", 0); SetTag("CurrentScreenManual", 0)
      Visibility <- "CurrentUserGroup"
   Button "Button_3" at 296,392 size 136x80; TextOff 'Statistici Productie'; Authorization "Monitor"
      on Press: ActivateScreen("Production.Repair", 0); SetTag("CurrentScreenStatistics", 0)
      Visibility <- "CurrentUserGroup"
   Button "Button_4" at 440,392 size 136x80; TextOff 'Alarme'; Authorization "Operate"
      on Press: ActivateScreen("Alarms", 0)
      Visibility <- "CurrentUserGroup"
   GraphicView "Graphic view_1" at 0,40 size 800x344; Picture "Vrancart V7 - cort-2"
   Group "Group" at 3,3 size 794x382
   GraphicIOField "Graphic I/O field_1" at 610,96 size 20x20; PictureList "List"
      ProcessValue <- "s_f{2}_step"
   GraphicIOField "Graphic I/O field_2" at 612,168 size 20x20; PictureList "List"
      ProcessValue <- "s_f{3}_step"
   GraphicIOField "Graphic I/O field_3" at 615,267 size 20x20; PictureList "List"
      ProcessValue <- "s_f{4}_step"
   GraphicIOField "Graphic I/O field_4" at 618,323 size 20x20; PictureList "List"
      ProcessValue <- "s_f{5}_step"
   GraphicIOField "Graphic I/O field_5" at 510,97 size 20x20; PictureList "List"
      ProcessValue <- "sn_f{1}_step"
   GraphicIOField "Graphic I/O field_6" at 512,169 size 20x20; PictureList "List"
      ProcessValue <- "sn_f{3}_step"
   GraphicIOField "Graphic I/O field_7" at 515,268 size 20x20; PictureList "List"
      ProcessValue <- "sn_f{4}_step"
   GraphicIOField "Graphic I/O field_8" at 518,324 size 20x20; PictureList "List"
      ProcessValue <- "sn_f{5}_step"
   GraphicView "Graphic view_10" at 129,149 size 15x15; Picture "Graphic_1"
      Visibility <- "Emergency Stop Destacker"
   GraphicView "Graphic view_11" at 511,62 size 15x15; Picture "Graphic_1"
      Visibility <- "Emergency Stop Zone 2"
   GraphicView "Graphic view_12" at 649,342 size 15x15; Picture "Graphic_1"
      Visibility <- "Emergency Stop Stacker"
   GraphicView "Graphic view_13" at 642,217 size 15x15; Picture "Graphic_1"
      Visibility <- "Stacker 115KF1 Safety Barrier Relay 2"
   GraphicView "Graphic view_14" at 584,211 size 15x15; Picture "Graphic_1"
      Visibility <- "Stacker 114KF1 Safety Barrier Relay 1"
   GraphicView "Graphic view_15" at 254,131 size 15x15; Picture "Graphic_1"
      Visibility <- "Destacker 111KF1 Safety Barrier Relay"
   Button "Button_9" at 558,40 size 96x32; TextOff '1200'
      on Press: SetBit("Length_S_HMI_1")
      Appearance <- "Fault_Length_S"
      Visibility <- "Fault_Length_S"
   Button "Button_10" at 558,95 size 96x32; TextOff '1600'
      on Press: SetBit("Length_S_HMI_2")
      Appearance <- "Fault_Length_S"
      Visibility <- "Fault_Length_S"
   Button "Button_11" at 558,150 size 96x32; TextOff '2000'
      on Press: SetBit("Length_S_HMI_3")
      Appearance <- "Fault_Length_S"
      Visibility <- "Fault_Length_S"
   Button "Button_12" at 558,205 size 96x32; TextOff 'OK'
      on Release: ResetBit("Fault_Length_DS_ACK")
      on Press: SetBit("Fault_Length_S_ACK")
      Visibility <- "Fault_Length_S"
   Button "Button_5" at 109,39 size 96x32; TextOff '1200'
      Appearance <- "Fault_Length_DS"
      on Press: SetBit("Length_DS_HMI_1")
      Visibility <- "Fault_Length_DS"
   Button "Button_6" at 109,94 size 96x32; TextOff '1600'
      Appearance <- "Fault_Length_DS"
      on Press: SetBit("Length_DS_HMI_2")
      Visibility <- "Fault_Length_DS"
   Button "Button_7" at 109,149 size 96x32; TextOff '2000'
      Appearance <- "Fault_Length_DS"
      on Press: SetBit("Length_DS_HMI_3")
      Visibility <- "Fault_Length_DS"
   Button "Button_8" at 109,204 size 96x32; TextOff 'OK'
      on Press: SetBit("Fault_Length_DS_ACK")
      on Release: ResetBit("Fault_Length_DS_ACK")
      Visibility <- "Fault_Length_DS"
   Line "Line_1" at 3,4 size 0x379
      Appearance <- "DB_MDM_SN_step"
   Line "Line_2" at 4,3 size 388x1
      Appearance <- "DB_MDM_SN_step"
   Line "Line_4" at 797,4 size 0x381
      Appearance <- "DB_MDM_S_step"
   Line "Line_5" at 394,4 size 400x0
      Appearance <- "DB_MDM_S_step"
   Line "Line_3" at 4,383 size 388x1
      Appearance <- "DB_MDM_SN_step"
   Line "Line_6" at 394,384 size 400x0
      Appearance <- "DB_MDM_S_step"
   GraphicView "Graphic view_2" at 610,96 size 20x20; Picture "Graphic_5"
      Visibility <- "s_f{2}_almt"
   GraphicView "Graphic view_3" at 612,168 size 20x20; Picture "Graphic_5"
      Visibility <- "s_f{3}_almt"
   GraphicView "Graphic view_4" at 615,267 size 20x20; Picture "Graphic_5"
      Visibility <- "s_f{4}_almt"
   GraphicView "Graphic view_5" at 618,323 size 20x20; Picture "Graphic_5"
      Visibility <- "s_f{5}_almt"
   GraphicView "Graphic view_6" at 510,97 size 20x20; Picture "Graphic_5"
      Visibility <- "sn_f{1}_almt"
   GraphicView "Graphic view_7" at 512,169 size 20x20; Picture "Graphic_5"
      Visibility <- "sn_f{3}_almt"
   GraphicView "Graphic view_8" at 515,268 size 20x20; Picture "Graphic_5"
      Visibility <- "sn_f{4}_almt"
   GraphicView "Graphic view_9" at 518,324 size 20x20; Picture "Graphic_5"
      Visibility <- "sn_f{5}_almt"

screen "Alarms" 800x480, template "TemplateWithClockAndBackBtn"
   AlarmView "Alarm view_1" at 0,40 size 800x348
   Button "Button_1" at 648,392 size 144x80; TextOff 'Confirmare Alarma Acknowledge'; Authorization "Operate"
      on Press: function_d9204949("Alarm view_1")
   Button "Button_2" at 8,392 size 144x80; TextOff 'Loguri Sistem / Acknowledge'; Authorization "Operate"
      on Press: ActivateScreen("SystemHealth", 0)

screen "SystemHealth" 800x480, template "TemplateWithClockAndBackBtn"
   SysDiagControl "System diagnostics view_1" at 0,40 size 800x440

screen "Settings" 800x480, template "TemplateWithClockAndBackBtn"
   UserView "User view_1" at 8,48 size 784x328
   Button "Button_1" at 8,392 size 96x80; TextOff 'Reset General'; Authorization "Operate"
   Button "Button_2" at 112,392 size 96x80; TextOff 'Reset Contoare'; Authorization "Operate"
   Button "Button_3" at 216,392 size 96x80; TextOff 'Calibrare Ecran'; Authorization "Operate"
      on Press: function_bc3e350c()
   Button "Button_4" at 320,392 size 96x80; TextOff 'Curatare Ecran'; Authorization "Operate"
      on Press: function_be740847(30)
   Button "Button_5" at 424,392 size 96x80; TextOff 'Stop Runtime'; Authorization "Operate"
      on Press: StopRuntime(0)

screen "Production.Repair" 800x480, template "TemplateWithClockAndBackBtnForStatistics"
   IOField "I/O field_1" at 696,48 size 96x32; FormatPattern 9
      ProcessValue <- "PalletsLastWeek"
   TextField "Text field_1" at 488,48 size 160x20; Text 'Paleti ultima saptamana'
   TextField "Text field_2" at 488,88 size 115x20; Text 'Paleti ultima luna'
   IOField "I/O field_2" at 696,88 size 96x32; FormatPattern 9
      ProcessValue <- "PalletsLastMonth"
   TrendView "Trend view_1" at 8,48 size 448x332
   IOField "I/O field_3" at 696,127 size 96x32; FormatPattern 99
      ProcessValue <- "DB20_DATA_HMI_Step_Destacker"
   TextField "Text field_3" at 488,127 size 97x20; Text 'Pas destivuire'
   TextField "Text field_4" at 488,167 size 81x20; Text 'Pas stivuire'
   IOField "I/O field_4" at 696,167 size 96x32; FormatPattern 99
      ProcessValue <- "DB20_DATA_HMI_Step_Stacker"
   Button "Button_1" at 488,256 size 124x97; TextOff 'REZ G7 DS'
      on Press: SetBit("Rez_G7_DS")
      on Release: ResetBit("Rez_G7_DS")
   Button "Button_2" at 650,256 size 124x97; TextOff 'REZ G7 S'
      on Press: SetBit("Rez_G7_S")
      on Release: ResetBit("Rez_G7_S")

screen "Production.Destroy" 800x480, template "TemplateWithClockAndBackBtnForStatistics"
   TrendView "Trend view_1" at 8,48 size 448x332

screen "Energy" 800x480, template "TemplateWithClockAndBackBtnForStatistics"
   IOField "I/O field_1" at 688,48 size 96x32; FormatPattern 9
      ProcessValue <- "FB_EnergyCounter_DB_Counters_LastHour_CV"
   TextField "Text field_3" at 600,48 size 70x20; Text 'Ultima ora'
   IOField "I/O field_2" at 688,88 size 96x32; FormatPattern 9
      ProcessValue <- "FB_EnergyCounter_DB_Counters_LastDay_CV"
   TextField "Text field_1" at 600,88 size 58x20; Text 'Ultima zi'
   IOField "I/O field_3" at 688,128 size 96x32; FormatPattern 9
      ProcessValue <- "FB_EnergyCounter_DB_Counters_LastMonth_CV"
   TextField "Text field_2" at 600,128 size 75x20; Text 'Ultima luna'
   TrendView "Trend view_1" at 8,48 size 448x332

screen "Safety" 800x480, template "TemplateWithClockAndBackBtnForStatistics"
   IOField "I/O field_1" at 336,48 size 96x32; FormatPattern 9
      ProcessValue <- "FB_AlarmCounter_DB_Counters_Destacker 110KF1 Safety Relay_CV"
   TextField "Text field_3" at 16,50 size 208x20; Text 'Destacker 110KF1 Safety Relay'
   IOField "I/O field_2" at 336,80 size 96x32; FormatPattern 9
      ProcessValue <- "FB_AlarmCounter_DB_Counters_Destacker 111KF1 Safety Barrier Relay_CV"
   TextField "Text field_1" at 16,82 size 257x20; Text 'Destacker 111KF1 Safety Barrier Relay'
   IOField "I/O field_3" at 336,112 size 96x32; FormatPattern 9
      ProcessValue <- "FB_AlarmCounter_DB_Counters_Zone 2 112KF1 Safety Relay_CV"
   TextField "Text field_2" at 16,114 size 185x20; Text 'Zone 2 112KF1 Safety Relay'
   IOField "I/O field_4" at 336,144 size 96x32; FormatPattern 9
      ProcessValue <- "FB_AlarmCounter_DB_Counters_Stacker 113KF1 Safety Relay_CV"
   TextField "Text field_4" at 16,146 size 192x20; Text 'Stacker 113KF1 Safety Relay'
   IOField "I/O field_5" at 336,176 size 96x32; FormatPattern 9
      ProcessValue <- "FB_AlarmCounter_DB_Counters_Stacker 114KF1 Safety Barrier Relay 1_CV"
   TextField "Text field_5" at 16,178 size 253x20; Text 'Stacker 114KF1 Safety Barrier Relay 1'
   IOField "I/O field_6" at 336,208 size 96x32; FormatPattern 9
      ProcessValue <- "FB_AlarmCounter_DB_Counters_Stacker 115KF1 Safety Barrier Relay 2_CV"
   TextField "Text field_6" at 16,210 size 253x20; Text 'Stacker 115KF1 Safety Barrier Relay 2'
   IOField "I/O field_7" at 336,240 size 96x32; FormatPattern 9
      ProcessValue <- "FB_AlarmCounter_DB_Counters_Emergency Stop Destacker_CV"
   TextField "Text field_7" at 16,242 size 180x20; Text 'Emergency Stop Destacker'
   IOField "I/O field_8" at 336,272 size 96x32; FormatPattern 9
      ProcessValue <- "FB_AlarmCounter_DB_Counters_Emergency Stop Zone 2_CV"
   TextField "Text field_8" at 16,274 size 157x20; Text 'Emergency Stop Zone 2'
   IOField "I/O field_9" at 336,304 size 96x32; FormatPattern 9
      ProcessValue <- "FB_AlarmCounter_DB_Counters_Emergency Stop Stacker_CV"
   TextField "Text field_9" at 16,306 size 164x20; Text 'Emergency Stop Stacker'
   Button "Button_1" at 552,160 size 128x64; TextOff 'Reset'; Authorization "User administration"

